REGION Network 7: IW272 - BWT Level (LT-422) - Tank #2
   RUNG wire#powerrail
      { S7_Templates := "[SrcType := Int, DestType := Real]" } Normalize(min := "20_TANKS_IP_DATA".RIO_04.SECOND_TANK.BWT_LEVEL_CNFG.RAW_MIN, value := "Tank 4S BWT Level", max := "20_TANKS_IP_DATA".RIO_04.SECOND_TANK.BWT_LEVEL_CNFG.RAW_MAX, out => "20_TANKS_IP_DATA".RIO_04.SECOND_TANK.BWT_LEVEL_CNFG.NORM)
      { S7_Templates := "[SrcType := Real, DestType := Real]" } Scale(min := "20_TANKS_IP_DATA".RIO_04.SECOND_TANK.BWT_LEVEL_CNFG.ENG_MIN, value := "IN_Level_WBT_4S", max := "20_TANKS_IP_DATA".RIO_04.SECOND_TANK.BWT_LEVEL_CNFG.ENG_MAX, out => "Tag_26")
      Move(in := "Data_From_WBT".Level_WBT_4S, out1 => "20_TANKS_IP_DATA".RIO_04.SECOND_TANK.BWT_LEVEL)
   END_RUNG
   // the same network as SCL:
   "20_TANKS_IP_DATA".RIO_04.SECOND_TANK.BWT_LEVEL_CNFG.NORM := NORM_X(MIN := "20_TANKS_IP_DATA".RIO_04.SECOND_TANK.BWT_LEVEL_CNFG.RAW_MIN, VALUE := "Tank 4S BWT Level", MAX := "20_TANKS_IP_DATA".RIO_04.SECOND_TANK.BWT_LEVEL_CNFG.RAW_MAX);
   "Tag_26" := SCALE_X(MIN := "20_TANKS_IP_DATA".RIO_04.SECOND_TANK.BWT_LEVEL_CNFG.ENG_MIN, VALUE := "IN_Level_WBT_4S", MAX := "20_TANKS_IP_DATA".RIO_04.SECOND_TANK.BWT_LEVEL_CNFG.ENG_MAX);
   "20_TANKS_IP_DATA".RIO_04.SECOND_TANK.BWT_LEVEL := "Data_From_WBT".Level_WBT_4S;
END_REGION

REGION Network 8: IW274 - Spare Input - Tank #1
   RUNG wire#powerrail
      { S7_Templates := "[SrcType := Int, DestType := Real]" } Normalize(min := "20_TANKS_IP_DATA".RIO_04.FIRST_TANK.SPARE_AI_1_CNFG.RAW_MIN, value := "RIO4_SPR_AI_274", max := "20_TANKS_IP_DATA".RIO_04.FIRST_TANK.SPARE_AI_1_CNFG.RAW_MAX, out => "20_TANKS_IP_DATA".RIO_04.FIRST_TANK.SPARE_AI_1_CNFG.NORM)
      { S7_Templates := "[SrcType := Real, DestType := Real]" } Scale(min := "20_TANKS_IP_DATA".RIO_04.FIRST_TANK.SPARE_AI_1_CNFG.ENG_MIN, value := "20_TANKS_IP_DATA".RIO_04.FIRST_TANK.SPARE_AI_1_CNFG.NORM, max := "20_TANKS_IP_DATA".RIO_04.FIRST_TANK.SPARE_AI_1_CNFG.ENG_MAX, out => "20_TANKS_IP_DATA".RIO_04.FIRST_TANK.SPARE_AI_1)
   END_RUNG
   // the same network as SCL:
   "20_TANKS_IP_DATA".RIO_04.FIRST_TANK.SPARE_AI_1_CNFG.NORM := NORM_X(MIN := "20_TANKS_IP_DATA".RIO_04.FIRST_TANK.SPARE_AI_1_CNFG.RAW_MIN, VALUE := "RIO4_SPR_AI_274", MAX := "20_TANKS_IP_DATA".RIO_04.FIRST_TANK.SPARE_AI_1_CNFG.RAW_MAX);
   "20_TANKS_IP_DATA".RIO_04.FIRST_TANK.SPARE_AI_1 := SCALE_X(MIN := "20_TANKS_IP_DATA".RIO_04.FIRST_TANK.SPARE_AI_1_CNFG.ENG_MIN, VALUE := "20_TANKS_IP_DATA".RIO_04.FIRST_TANK.SPARE_AI_1_CNFG.NORM, MAX := "20_TANKS_IP_DATA".RIO_04.FIRST_TANK.SPARE_AI_1_CNFG.ENG_MAX);
END_REGION

REGION Network 9: IW276 - BWT Ph (426) - Tank #1
   RUNG wire#powerrail
      { S7_Templates := "[SrcType := Int, DestType := Real]" } Normalize(min := "20_TANKS_IP_DATA".RIO_04.FIRST_TANK.BWT_PH_CNFG.RAW_MIN, value := "Tank 4P BWT ph", max := "20_TANKS_IP_DATA".RIO_04.FIRST_TANK.BWT_PH_CNFG.RAW_MAX, out => "20_TANKS_IP_DATA".RIO_04.FIRST_TANK.BWT_PH_CNFG.NORM)
      { S7_Templates := "[SrcType := Real, DestType := Real]" } Scale(min := "20_TANKS_IP_DATA".RIO_04.FIRST_TANK.BWT_PH_CNFG.ENG_MIN, value := "20_TANKS_IP_DATA".RIO_04.FIRST_TANK.BWT_PH_CNFG.NORM, max := "20_TANKS_IP_DATA".RIO_04.FIRST_TANK.BWT_PH_CNFG.ENG_MAX, out => "20_TANKS_IP_DATA".RIO_04.FIRST_TANK.BWT_PH)
   END_RUNG
   // the same network as SCL:
   "20_TANKS_IP_DATA".RIO_04.FIRST_TANK.BWT_PH_CNFG.NORM := NORM_X(MIN := "20_TANKS_IP_DATA".RIO_04.FIRST_TANK.BWT_PH_CNFG.RAW_MIN, VALUE := "Tank 4P BWT ph", MAX := "20_TANKS_IP_DATA".RIO_04.FIRST_TANK.BWT_PH_CNFG.RAW_MAX);
   "20_TANKS_IP_DATA".RIO_04.FIRST_TANK.BWT_PH := SCALE_X(MIN := "20_TANKS_IP_DATA".RIO_04.FIRST_TANK.BWT_PH_CNFG.ENG_MIN, VALUE := "20_TANKS_IP_DATA".RIO_04.FIRST_TANK.BWT_PH_CNFG.NORM, MAX := "20_TANKS_IP_DATA".RIO_04.FIRST_TANK.BWT_PH_CNFG.ENG_MAX);
END_REGION

REGION Network 10: IW278 - BWT Temperature (426) - Tank #1
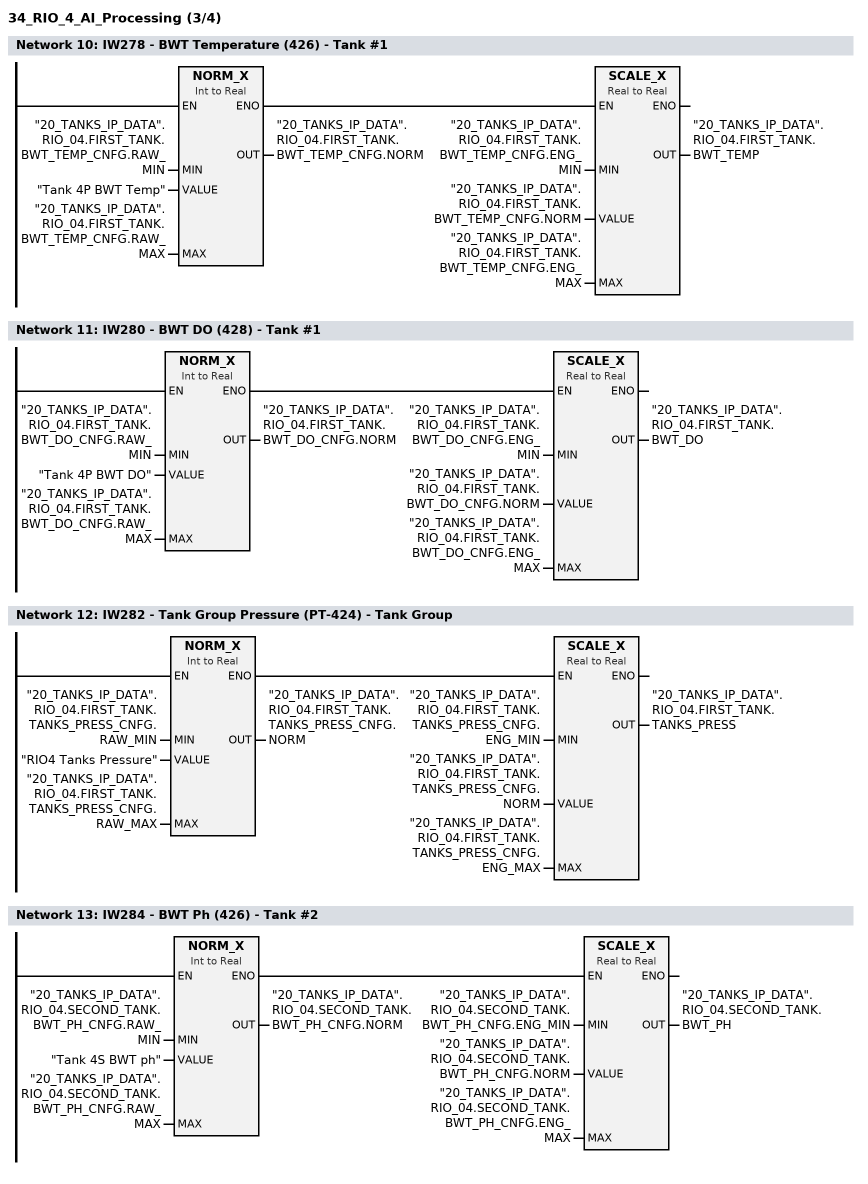
   RUNG wire#powerrail
      { S7_Templates := "[SrcType := Int, DestType := Real]" } Normalize(min := "20_TANKS_IP_DATA".RIO_04.FIRST_TANK.BWT_TEMP_CNFG.RAW_MIN, value := "Tank 4P BWT Temp", max := "20_TANKS_IP_DATA".RIO_04.FIRST_TANK.BWT_TEMP_CNFG.RAW_MAX, out => "20_TANKS_IP_DATA".RIO_04.FIRST_TANK.BWT_TEMP_CNFG.NORM)
      { S7_Templates := "[SrcType := Real, DestType := Real]" } Scale(min := "20_TANKS_IP_DATA".RIO_04.FIRST_TANK.BWT_TEMP_CNFG.ENG_MIN, value := "20_TANKS_IP_DATA".RIO_04.FIRST_TANK.BWT_TEMP_CNFG.NORM, max := "20_TANKS_IP_DATA".RIO_04.FIRST_TANK.BWT_TEMP_CNFG.ENG_MAX, out => "20_TANKS_IP_DATA".RIO_04.FIRST_TANK.BWT_TEMP)
   END_RUNG
   // the same network as SCL:
   "20_TANKS_IP_DATA".RIO_04.FIRST_TANK.BWT_TEMP_CNFG.NORM := NORM_X(MIN := "20_TANKS_IP_DATA".RIO_04.FIRST_TANK.BWT_TEMP_CNFG.RAW_MIN, VALUE := "Tank 4P BWT Temp", MAX := "20_TANKS_IP_DATA".RIO_04.FIRST_TANK.BWT_TEMP_CNFG.RAW_MAX);
   "20_TANKS_IP_DATA".RIO_04.FIRST_TANK.BWT_TEMP := SCALE_X(MIN := "20_TANKS_IP_DATA".RIO_04.FIRST_TANK.BWT_TEMP_CNFG.ENG_MIN, VALUE := "20_TANKS_IP_DATA".RIO_04.FIRST_TANK.BWT_TEMP_CNFG.NORM, MAX := "20_TANKS_IP_DATA".RIO_04.FIRST_TANK.BWT_TEMP_CNFG.ENG_MAX);
END_REGION

REGION Network 11: IW280 - BWT DO (428) - Tank #1
   RUNG wire#powerrail
      { S7_Templates := "[SrcType := Int, DestType := Real]" } Normalize(min := "20_TANKS_IP_DATA".RIO_04.FIRST_TANK.BWT_DO_CNFG.RAW_MIN, value := "Tank 4P BWT DO", max := "20_TANKS_IP_DATA".RIO_04.FIRST_TANK.BWT_DO_CNFG.RAW_MAX, out => "20_TANKS_IP_DATA".RIO_04.FIRST_TANK.BWT_DO_CNFG.NORM)
      { S7_Templates := "[SrcType := Real, DestType := Real]" } Scale(min := "20_TANKS_IP_DATA".RIO_04.FIRST_TANK.BWT_DO_CNFG.ENG_MIN, value := "20_TANKS_IP_DATA".RIO_04.FIRST_TANK.BWT_DO_CNFG.NORM, max := "20_TANKS_IP_DATA".RIO_04.FIRST_TANK.BWT_DO_CNFG.ENG_MAX, out => "20_TANKS_IP_DATA".RIO_04.FIRST_TANK.BWT_DO)
   END_RUNG
   // the same network as SCL:
   "20_TANKS_IP_DATA".RIO_04.FIRST_TANK.BWT_DO_CNFG.NORM := NORM_X(MIN := "20_TANKS_IP_DATA".RIO_04.FIRST_TANK.BWT_DO_CNFG.RAW_MIN, VALUE := "Tank 4P BWT DO", MAX := "20_TANKS_IP_DATA".RIO_04.FIRST_TANK.BWT_DO_CNFG.RAW_MAX);
   "20_TANKS_IP_DATA".RIO_04.FIRST_TANK.BWT_DO := SCALE_X(MIN := "20_TANKS_IP_DATA".RIO_04.FIRST_TANK.BWT_DO_CNFG.ENG_MIN, VALUE := "20_TANKS_IP_DATA".RIO_04.FIRST_TANK.BWT_DO_CNFG.NORM, MAX := "20_TANKS_IP_DATA".RIO_04.FIRST_TANK.BWT_DO_CNFG.ENG_MAX);
END_REGION

REGION Network 12: IW282 - Tank Group Pressure (PT-424) - Tank Group
   RUNG wire#powerrail
      { S7_Templates := "[SrcType := Int, DestType := Real]" } Normalize(min := "20_TANKS_IP_DATA".RIO_04.FIRST_TANK.TANKS_PRESS_CNFG.RAW_MIN, value := "RIO4 Tanks Pressure", max := "20_TANKS_IP_DATA".RIO_04.FIRST_TANK.TANKS_PRESS_CNFG.RAW_MAX, out => "20_TANKS_IP_DATA".RIO_04.FIRST_TANK.TANKS_PRESS_CNFG.NORM)
      { S7_Templates := "[SrcType := Real, DestType := Real]" } Scale(min := "20_TANKS_IP_DATA".RIO_04.FIRST_TANK.TANKS_PRESS_CNFG.ENG_MIN, value := "20_TANKS_IP_DATA".RIO_04.FIRST_TANK.TANKS_PRESS_CNFG.NORM, max := "20_TANKS_IP_DATA".RIO_04.FIRST_TANK.TANKS_PRESS_CNFG.ENG_MAX, out => "20_TANKS_IP_DATA".RIO_04.FIRST_TANK.TANKS_PRESS)
   END_RUNG
   // the same network as SCL:
   "20_TANKS_IP_DATA".RIO_04.FIRST_TANK.TANKS_PRESS_CNFG.NORM := NORM_X(MIN := "20_TANKS_IP_DATA".RIO_04.FIRST_TANK.TANKS_PRESS_CNFG.RAW_MIN, VALUE := "RIO4 Tanks Pressure", MAX := "20_TANKS_IP_DATA".RIO_04.FIRST_TANK.TANKS_PRESS_CNFG.RAW_MAX);
   "20_TANKS_IP_DATA".RIO_04.FIRST_TANK.TANKS_PRESS := SCALE_X(MIN := "20_TANKS_IP_DATA".RIO_04.FIRST_TANK.TANKS_PRESS_CNFG.ENG_MIN, VALUE := "20_TANKS_IP_DATA".RIO_04.FIRST_TANK.TANKS_PRESS_CNFG.NORM, MAX := "20_TANKS_IP_DATA".RIO_04.FIRST_TANK.TANKS_PRESS_CNFG.ENG_MAX);
END_REGION

REGION Network 13: IW284 - BWT Ph (426) - Tank #2
   RUNG wire#powerrail
      { S7_Templates := "[SrcType := Int, DestType := Real]" } Normalize(min := "20_TANKS_IP_DATA".RIO_04.SECOND_TANK.BWT_PH_CNFG.RAW_MIN, value := "Tank 4S BWT ph", max := "20_TANKS_IP_DATA".RIO_04.SECOND_TANK.BWT_PH_CNFG.RAW_MAX, out => "20_TANKS_IP_DATA".RIO_04.SECOND_TANK.BWT_PH_CNFG.NORM)
      { S7_Templates := "[SrcType := Real, DestType := Real]" } Scale(min := "20_TANKS_IP_DATA".RIO_04.SECOND_TANK.BWT_PH_CNFG.ENG_MIN, value := "20_TANKS_IP_DATA".RIO_04.SECOND_TANK.BWT_PH_CNFG.NORM, max := "20_TANKS_IP_DATA".RIO_04.SECOND_TANK.BWT_PH_CNFG.ENG_MAX, out => "20_TANKS_IP_DATA".RIO_04.SECOND_TANK.BWT_PH)
   END_RUNG
   // the same network as SCL:
   "20_TANKS_IP_DATA".RIO_04.SECOND_TANK.BWT_PH_CNFG.NORM := NORM_X(MIN := "20_TANKS_IP_DATA".RIO_04.SECOND_TANK.BWT_PH_CNFG.RAW_MIN, VALUE := "Tank 4S BWT ph", MAX := "20_TANKS_IP_DATA".RIO_04.SECOND_TANK.BWT_PH_CNFG.RAW_MAX);
   "20_TANKS_IP_DATA".RIO_04.SECOND_TANK.BWT_PH := SCALE_X(MIN := "20_TANKS_IP_DATA".RIO_04.SECOND_TANK.BWT_PH_CNFG.ENG_MIN, VALUE := "20_TANKS_IP_DATA".RIO_04.SECOND_TANK.BWT_PH_CNFG.NORM, MAX := "20_TANKS_IP_DATA".RIO_04.SECOND_TANK.BWT_PH_CNFG.ENG_MAX);
END_REGION

REGION Network 14: IW286 - BWT Temperature (426) - Tank #2
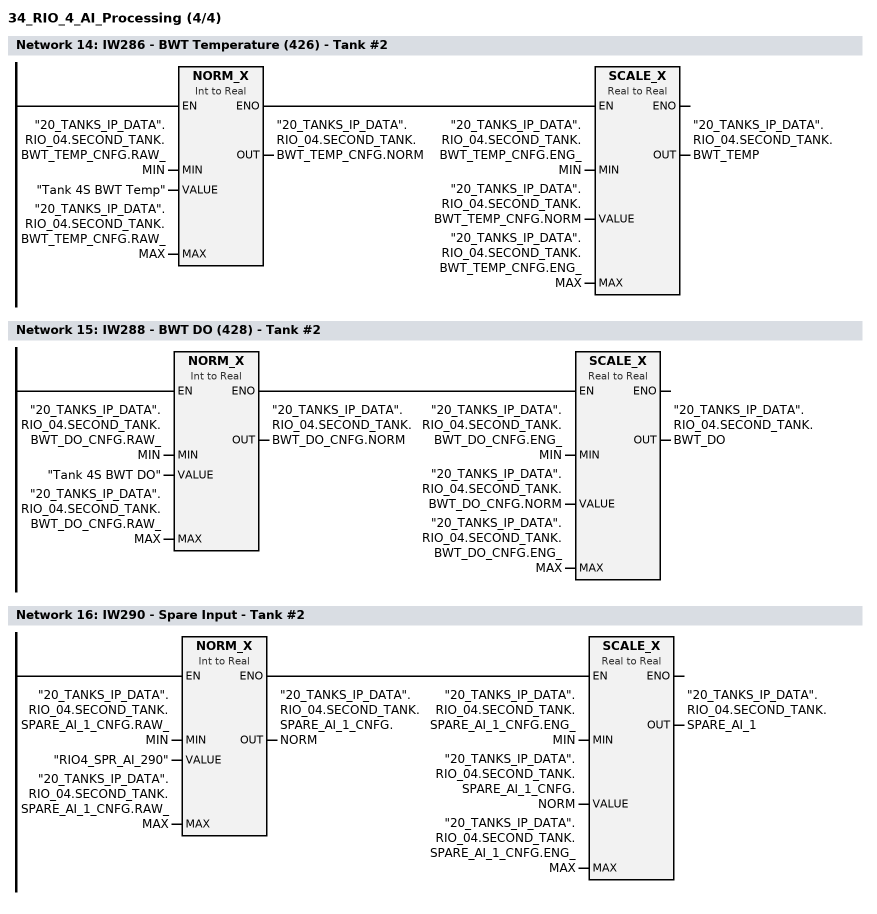
   RUNG wire#powerrail
      { S7_Templates := "[SrcType := Int, DestType := Real]" } Normalize(min := "20_TANKS_IP_DATA".RIO_04.SECOND_TANK.BWT_TEMP_CNFG.RAW_MIN, value := "Tank 4S BWT Temp", max := "20_TANKS_IP_DATA".RIO_04.SECOND_TANK.BWT_TEMP_CNFG.RAW_MAX, out => "20_TANKS_IP_DATA".RIO_04.SECOND_TANK.BWT_TEMP_CNFG.NORM)
      { S7_Templates := "[SrcType := Real, DestType := Real]" } Scale(min := "20_TANKS_IP_DATA".RIO_04.SECOND_TANK.BWT_TEMP_CNFG.ENG_MIN, value := "20_TANKS_IP_DATA".RIO_04.SECOND_TANK.BWT_TEMP_CNFG.NORM, max := "20_TANKS_IP_DATA".RIO_04.SECOND_TANK.BWT_TEMP_CNFG.ENG_MAX, out => "20_TANKS_IP_DATA".RIO_04.SECOND_TANK.BWT_TEMP)
   END_RUNG
   // the same network as SCL:
   "20_TANKS_IP_DATA".RIO_04.SECOND_TANK.BWT_TEMP_CNFG.NORM := NORM_X(MIN := "20_TANKS_IP_DATA".RIO_04.SECOND_TANK.BWT_TEMP_CNFG.RAW_MIN, VALUE := "Tank 4S BWT Temp", MAX := "20_TANKS_IP_DATA".RIO_04.SECOND_TANK.BWT_TEMP_CNFG.RAW_MAX);
   "20_TANKS_IP_DATA".RIO_04.SECOND_TANK.BWT_TEMP := SCALE_X(MIN := "20_TANKS_IP_DATA".RIO_04.SECOND_TANK.BWT_TEMP_CNFG.ENG_MIN, VALUE := "20_TANKS_IP_DATA".RIO_04.SECOND_TANK.BWT_TEMP_CNFG.NORM, MAX := "20_TANKS_IP_DATA".RIO_04.SECOND_TANK.BWT_TEMP_CNFG.ENG_MAX);
END_REGION

REGION Network 15: IW288 - BWT DO (428) - Tank #2
   RUNG wire#powerrail
      { S7_Templates := "[SrcType := Int, DestType := Real]" } Normalize(min := "20_TANKS_IP_DATA".RIO_04.SECOND_TANK.BWT_DO_CNFG.RAW_MIN, value := "Tank 4S BWT DO", max := "20_TANKS_IP_DATA".RIO_04.SECOND_TANK.BWT_DO_CNFG.RAW_MAX, out => "20_TANKS_IP_DATA".RIO_04.SECOND_TANK.BWT_DO_CNFG.NORM)
      { S7_Templates := "[SrcType := Real, DestType := Real]" } Scale(min := "20_TANKS_IP_DATA".RIO_04.SECOND_TANK.BWT_DO_CNFG.ENG_MIN, value := "20_TANKS_IP_DATA".RIO_04.SECOND_TANK.BWT_DO_CNFG.NORM, max := "20_TANKS_IP_DATA".RIO_04.SECOND_TANK.BWT_DO_CNFG.ENG_MAX, out => "20_TANKS_IP_DATA".RIO_04.SECOND_TANK.BWT_DO)
   END_RUNG
   // the same network as SCL:
   "20_TANKS_IP_DATA".RIO_04.SECOND_TANK.BWT_DO_CNFG.NORM := NORM_X(MIN := "20_TANKS_IP_DATA".RIO_04.SECOND_TANK.BWT_DO_CNFG.RAW_MIN, VALUE := "Tank 4S BWT DO", MAX := "20_TANKS_IP_DATA".RIO_04.SECOND_TANK.BWT_DO_CNFG.RAW_MAX);
   "20_TANKS_IP_DATA".RIO_04.SECOND_TANK.BWT_DO := SCALE_X(MIN := "20_TANKS_IP_DATA".RIO_04.SECOND_TANK.BWT_DO_CNFG.ENG_MIN, VALUE := "20_TANKS_IP_DATA".RIO_04.SECOND_TANK.BWT_DO_CNFG.NORM, MAX := "20_TANKS_IP_DATA".RIO_04.SECOND_TANK.BWT_DO_CNFG.ENG_MAX);
END_REGION

REGION Network 16: IW290 - Spare Input - Tank #2
   RUNG wire#powerrail
      { S7_Templates := "[SrcType := Int, DestType := Real]" } Normalize(min := "20_TANKS_IP_DATA".RIO_04.SECOND_TANK.SPARE_AI_1_CNFG.RAW_MIN, value := "RIO4_SPR_AI_290", max := "20_TANKS_IP_DATA".RIO_04.SECOND_TANK.SPARE_AI_1_CNFG.RAW_MAX, out => "20_TANKS_IP_DATA".RIO_04.SECOND_TANK.SPARE_AI_1_CNFG.NORM)
      { S7_Templates := "[SrcType := Real, DestType := Real]" } Scale(min := "20_TANKS_IP_DATA".RIO_04.SECOND_TANK.SPARE_AI_1_CNFG.ENG_MIN, value := "20_TANKS_IP_DATA".RIO_04.SECOND_TANK.SPARE_AI_1_CNFG.NORM, max := "20_TANKS_IP_DATA".RIO_04.SECOND_TANK.SPARE_AI_1_CNFG.ENG_MAX, out => "20_TANKS_IP_DATA".RIO_04.SECOND_TANK.SPARE_AI_1)
   END_RUNG
   // the same network as SCL:
   "20_TANKS_IP_DATA".RIO_04.SECOND_TANK.SPARE_AI_1_CNFG.NORM := NORM_X(MIN := "20_TANKS_IP_DATA".RIO_04.SECOND_TANK.SPARE_AI_1_CNFG.RAW_MIN, VALUE := "RIO4_SPR_AI_290", MAX := "20_TANKS_IP_DATA".RIO_04.SECOND_TANK.SPARE_AI_1_CNFG.RAW_MAX);
   "20_TANKS_IP_DATA".RIO_04.SECOND_TANK.SPARE_AI_1 := SCALE_X(MIN := "20_TANKS_IP_DATA".RIO_04.SECOND_TANK.SPARE_AI_1_CNFG.ENG_MIN, VALUE := "20_TANKS_IP_DATA".RIO_04.SECOND_TANK.SPARE_AI_1_CNFG.NORM, MAX := "20_TANKS_IP_DATA".RIO_04.SECOND_TANK.SPARE_AI_1_CNFG.ENG_MAX);
END_REGION
END_FUNCTION

FUNCTION "35_RIO_5_AI_Processing" : Void   // FC35, LAD
TITLE = Analogue Input Processing (Tank 1 = 5P, Tank 2 = 5S)
{ S7_Optimized_Access := 'TRUE' }
AUTHOR : JRS
VERSION : 0.1
// To process raw inputs prior to code use
BEGIN

REGION Network 1: IW300 - USD Flow (FIT-418) - Tank #1
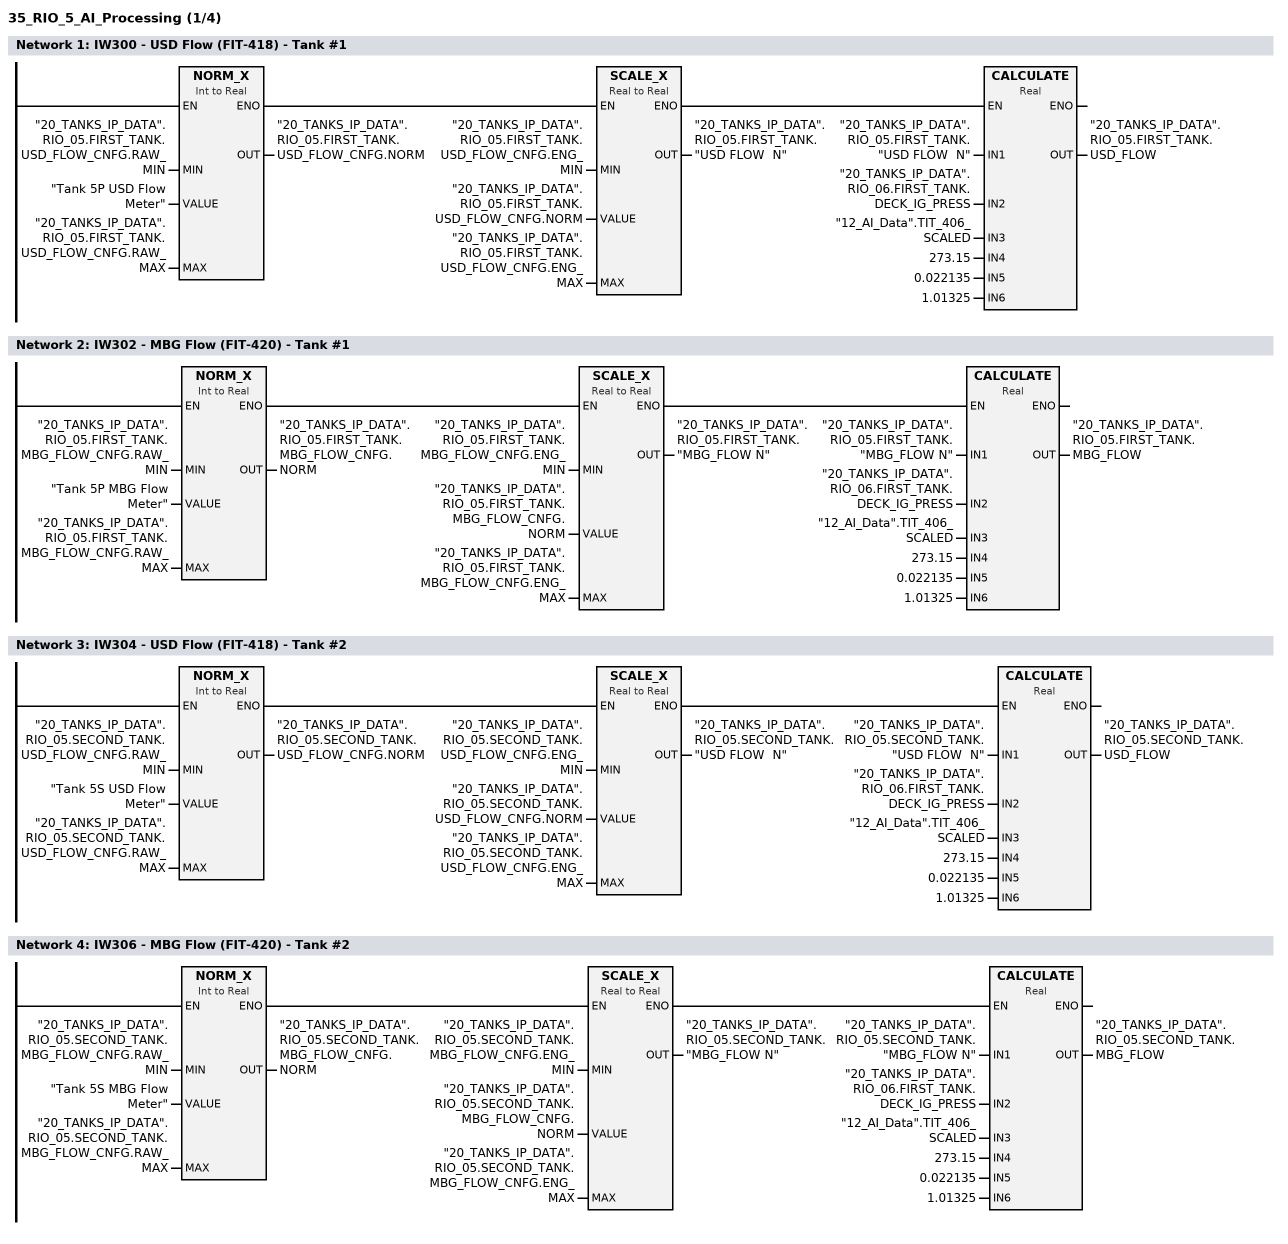
   RUNG wire#powerrail
      { S7_Templates := "[SrcType := Int, DestType := Real]" } Normalize(min := "20_TANKS_IP_DATA".RIO_05.FIRST_TANK.USD_FLOW_CNFG.RAW_MIN, value := "Tank 5P USD Flow Meter", max := "20_TANKS_IP_DATA".RIO_05.FIRST_TANK.USD_FLOW_CNFG.RAW_MAX, out => "20_TANKS_IP_DATA".RIO_05.FIRST_TANK.USD_FLOW_CNFG.NORM)
      { S7_Templates := "[SrcType := Real, DestType := Real]" } Scale(min := "20_TANKS_IP_DATA".RIO_05.FIRST_TANK.USD_FLOW_CNFG.ENG_MIN, value := "20_TANKS_IP_DATA".RIO_05.FIRST_TANK.USD_FLOW_CNFG.NORM, max := "20_TANKS_IP_DATA".RIO_05.FIRST_TANK.USD_FLOW_CNFG.ENG_MAX, out => "20_TANKS_IP_DATA".RIO_05.FIRST_TANK."USD FLOW  N")
      { S7_Templates := "SrcType := Real"; S7_Expression := "IN1*(IN2+IN6)/IN6*IN4/(IN3+IN4)" } Calculate(in1 := "20_TANKS_IP_DATA".RIO_05.FIRST_TANK."USD FLOW  N", in2 := "20_TANKS_IP_DATA".RIO_06.FIRST_TANK.DECK_IG_PRESS, in3 := "12_AI_Data".TIT_406_SCALED, in4 := 273.15, in5 := 0.022135, in6 := 1.01325, out => "20_TANKS_IP_DATA".RIO_05.FIRST_TANK.USD_FLOW)
   END_RUNG
   // the same network as SCL:
   "20_TANKS_IP_DATA".RIO_05.FIRST_TANK.USD_FLOW_CNFG.NORM := NORM_X(MIN := "20_TANKS_IP_DATA".RIO_05.FIRST_TANK.USD_FLOW_CNFG.RAW_MIN, VALUE := "Tank 5P USD Flow Meter", MAX := "20_TANKS_IP_DATA".RIO_05.FIRST_TANK.USD_FLOW_CNFG.RAW_MAX);
   "20_TANKS_IP_DATA".RIO_05.FIRST_TANK."USD FLOW  N" := SCALE_X(MIN := "20_TANKS_IP_DATA".RIO_05.FIRST_TANK.USD_FLOW_CNFG.ENG_MIN, VALUE := "20_TANKS_IP_DATA".RIO_05.FIRST_TANK.USD_FLOW_CNFG.NORM, MAX := "20_TANKS_IP_DATA".RIO_05.FIRST_TANK.USD_FLOW_CNFG.ENG_MAX);
   "20_TANKS_IP_DATA".RIO_05.FIRST_TANK.USD_FLOW := "20_TANKS_IP_DATA".RIO_05.FIRST_TANK."USD FLOW  N"*("20_TANKS_IP_DATA".RIO_06.FIRST_TANK.DECK_IG_PRESS+1.01325)/1.01325*273.15/("12_AI_Data".TIT_406_SCALED+273.15);
END_REGION

REGION Network 2: IW302 - MBG Flow (FIT-420) - Tank #1
   RUNG wire#powerrail
      { S7_Templates := "[SrcType := Int, DestType := Real]" } Normalize(min := "20_TANKS_IP_DATA".RIO_05.FIRST_TANK.MBG_FLOW_CNFG.RAW_MIN, value := "Tank 5P MBG Flow Meter", max := "20_TANKS_IP_DATA".RIO_05.FIRST_TANK.MBG_FLOW_CNFG.RAW_MAX, out => "20_TANKS_IP_DATA".RIO_05.FIRST_TANK.MBG_FLOW_CNFG.NORM)
      { S7_Templates := "[SrcType := Real, DestType := Real]" } Scale(min := "20_TANKS_IP_DATA".RIO_05.FIRST_TANK.MBG_FLOW_CNFG.ENG_MIN, value := "20_TANKS_IP_DATA".RIO_05.FIRST_TANK.MBG_FLOW_CNFG.NORM, max := "20_TANKS_IP_DATA".RIO_05.FIRST_TANK.MBG_FLOW_CNFG.ENG_MAX, out => "20_TANKS_IP_DATA".RIO_05.FIRST_TANK."MBG_FLOW N")
      { S7_Templates := "SrcType := Real"; S7_Expression := "IN1*(IN2+IN6)/IN6*IN4/(IN3+IN4)" } Calculate(in1 := "20_TANKS_IP_DATA".RIO_05.FIRST_TANK."MBG_FLOW N", in2 := "20_TANKS_IP_DATA".RIO_06.FIRST_TANK.DECK_IG_PRESS, in3 := "12_AI_Data".TIT_406_SCALED, in4 := 273.15, in5 := 0.022135, in6 := 1.01325, out => "20_TANKS_IP_DATA".RIO_05.FIRST_TANK.MBG_FLOW)
   END_RUNG
   // the same network as SCL:
   "20_TANKS_IP_DATA".RIO_05.FIRST_TANK.MBG_FLOW_CNFG.NORM := NORM_X(MIN := "20_TANKS_IP_DATA".RIO_05.FIRST_TANK.MBG_FLOW_CNFG.RAW_MIN, VALUE := "Tank 5P MBG Flow Meter", MAX := "20_TANKS_IP_DATA".RIO_05.FIRST_TANK.MBG_FLOW_CNFG.RAW_MAX);
   "20_TANKS_IP_DATA".RIO_05.FIRST_TANK."MBG_FLOW N" := SCALE_X(MIN := "20_TANKS_IP_DATA".RIO_05.FIRST_TANK.MBG_FLOW_CNFG.ENG_MIN, VALUE := "20_TANKS_IP_DATA".RIO_05.FIRST_TANK.MBG_FLOW_CNFG.NORM, MAX := "20_TANKS_IP_DATA".RIO_05.FIRST_TANK.MBG_FLOW_CNFG.ENG_MAX);
   "20_TANKS_IP_DATA".RIO_05.FIRST_TANK.MBG_FLOW := "20_TANKS_IP_DATA".RIO_05.FIRST_TANK."MBG_FLOW N"*("20_TANKS_IP_DATA".RIO_06.FIRST_TANK.DECK_IG_PRESS+1.01325)/1.01325*273.15/("12_AI_Data".TIT_406_SCALED+273.15);
END_REGION

REGION Network 3: IW304 - USD Flow (FIT-418) - Tank #2
   RUNG wire#powerrail
      { S7_Templates := "[SrcType := Int, DestType := Real]" } Normalize(min := "20_TANKS_IP_DATA".RIO_05.SECOND_TANK.USD_FLOW_CNFG.RAW_MIN, value := "Tank 5S USD Flow Meter", max := "20_TANKS_IP_DATA".RIO_05.SECOND_TANK.USD_FLOW_CNFG.RAW_MAX, out => "20_TANKS_IP_DATA".RIO_05.SECOND_TANK.USD_FLOW_CNFG.NORM)
      { S7_Templates := "[SrcType := Real, DestType := Real]" } Scale(min := "20_TANKS_IP_DATA".RIO_05.SECOND_TANK.USD_FLOW_CNFG.ENG_MIN, value := "20_TANKS_IP_DATA".RIO_05.SECOND_TANK.USD_FLOW_CNFG.NORM, max := "20_TANKS_IP_DATA".RIO_05.SECOND_TANK.USD_FLOW_CNFG.ENG_MAX, out => "20_TANKS_IP_DATA".RIO_05.SECOND_TANK."USD FLOW  N")
      { S7_Templates := "SrcType := Real"; S7_Expression := "IN1*(IN2+IN6)/IN6*IN4/(IN3+IN4)" } Calculate(in1 := "20_TANKS_IP_DATA".RIO_05.SECOND_TANK."USD FLOW  N", in2 := "20_TANKS_IP_DATA".RIO_06.FIRST_TANK.DECK_IG_PRESS, in3 := "12_AI_Data".TIT_406_SCALED, in4 := 273.15, in5 := 0.022135, in6 := 1.01325, out => "20_TANKS_IP_DATA".RIO_05.SECOND_TANK.USD_FLOW)
   END_RUNG
   // the same network as SCL:
   "20_TANKS_IP_DATA".RIO_05.SECOND_TANK.USD_FLOW_CNFG.NORM := NORM_X(MIN := "20_TANKS_IP_DATA".RIO_05.SECOND_TANK.USD_FLOW_CNFG.RAW_MIN, VALUE := "Tank 5S USD Flow Meter", MAX := "20_TANKS_IP_DATA".RIO_05.SECOND_TANK.USD_FLOW_CNFG.RAW_MAX);
   "20_TANKS_IP_DATA".RIO_05.SECOND_TANK."USD FLOW  N" := SCALE_X(MIN := "20_TANKS_IP_DATA".RIO_05.SECOND_TANK.USD_FLOW_CNFG.ENG_MIN, VALUE := "20_TANKS_IP_DATA".RIO_05.SECOND_TANK.USD_FLOW_CNFG.NORM, MAX := "20_TANKS_IP_DATA".RIO_05.SECOND_TANK.USD_FLOW_CNFG.ENG_MAX);
   "20_TANKS_IP_DATA".RIO_05.SECOND_TANK.USD_FLOW := "20_TANKS_IP_DATA".RIO_05.SECOND_TANK."USD FLOW  N"*("20_TANKS_IP_DATA".RIO_06.FIRST_TANK.DECK_IG_PRESS+1.01325)/1.01325*273.15/("12_AI_Data".TIT_406_SCALED+273.15);
END_REGION

REGION Network 4: IW306 - MBG Flow (FIT-420) - Tank #2
   RUNG wire#powerrail
      { S7_Templates := "[SrcType := Int, DestType := Real]" } Normalize(min := "20_TANKS_IP_DATA".RIO_05.SECOND_TANK.MBG_FLOW_CNFG.RAW_MIN, value := "Tank 5S MBG Flow Meter", max := "20_TANKS_IP_DATA".RIO_05.SECOND_TANK.MBG_FLOW_CNFG.RAW_MAX, out => "20_TANKS_IP_DATA".RIO_05.SECOND_TANK.MBG_FLOW_CNFG.NORM)
      { S7_Templates := "[SrcType := Real, DestType := Real]" } Scale(min := "20_TANKS_IP_DATA".RIO_05.SECOND_TANK.MBG_FLOW_CNFG.ENG_MIN, value := "20_TANKS_IP_DATA".RIO_05.SECOND_TANK.MBG_FLOW_CNFG.NORM, max := "20_TANKS_IP_DATA".RIO_05.SECOND_TANK.MBG_FLOW_CNFG.ENG_MAX, out => "20_TANKS_IP_DATA".RIO_05.SECOND_TANK."MBG_FLOW N")
      { S7_Templates := "SrcType := Real"; S7_Expression := "IN1*(IN2+IN6)/IN6*IN4/(IN3+IN4)" } Calculate(in1 := "20_TANKS_IP_DATA".RIO_05.SECOND_TANK."MBG_FLOW N", in2 := "20_TANKS_IP_DATA".RIO_06.FIRST_TANK.DECK_IG_PRESS, in3 := "12_AI_Data".TIT_406_SCALED, in4 := 273.15, in5 := 0.022135, in6 := 1.01325, out => "20_TANKS_IP_DATA".RIO_05.SECOND_TANK.MBG_FLOW)
   END_RUNG
   // the same network as SCL:
   "20_TANKS_IP_DATA".RIO_05.SECOND_TANK.MBG_FLOW_CNFG.NORM := NORM_X(MIN := "20_TANKS_IP_DATA".RIO_05.SECOND_TANK.MBG_FLOW_CNFG.RAW_MIN, VALUE := "Tank 5S MBG Flow Meter", MAX := "20_TANKS_IP_DATA".RIO_05.SECOND_TANK.MBG_FLOW_CNFG.RAW_MAX);
   "20_TANKS_IP_DATA".RIO_05.SECOND_TANK."MBG_FLOW N" := SCALE_X(MIN := "20_TANKS_IP_DATA".RIO_05.SECOND_TANK.MBG_FLOW_CNFG.ENG_MIN, VALUE := "20_TANKS_IP_DATA".RIO_05.SECOND_TANK.MBG_FLOW_CNFG.NORM, MAX := "20_TANKS_IP_DATA".RIO_05.SECOND_TANK.MBG_FLOW_CNFG.ENG_MAX);
   "20_TANKS_IP_DATA".RIO_05.SECOND_TANK.MBG_FLOW := "20_TANKS_IP_DATA".RIO_05.SECOND_TANK."MBG_FLOW N"*("20_TANKS_IP_DATA".RIO_06.FIRST_TANK.DECK_IG_PRESS+1.01325)/1.01325*273.15/("12_AI_Data".TIT_406_SCALED+273.15);
END_REGION

REGION Network 5: IW308 - Deck Main IG Pressure (PT-415) - Tank Group
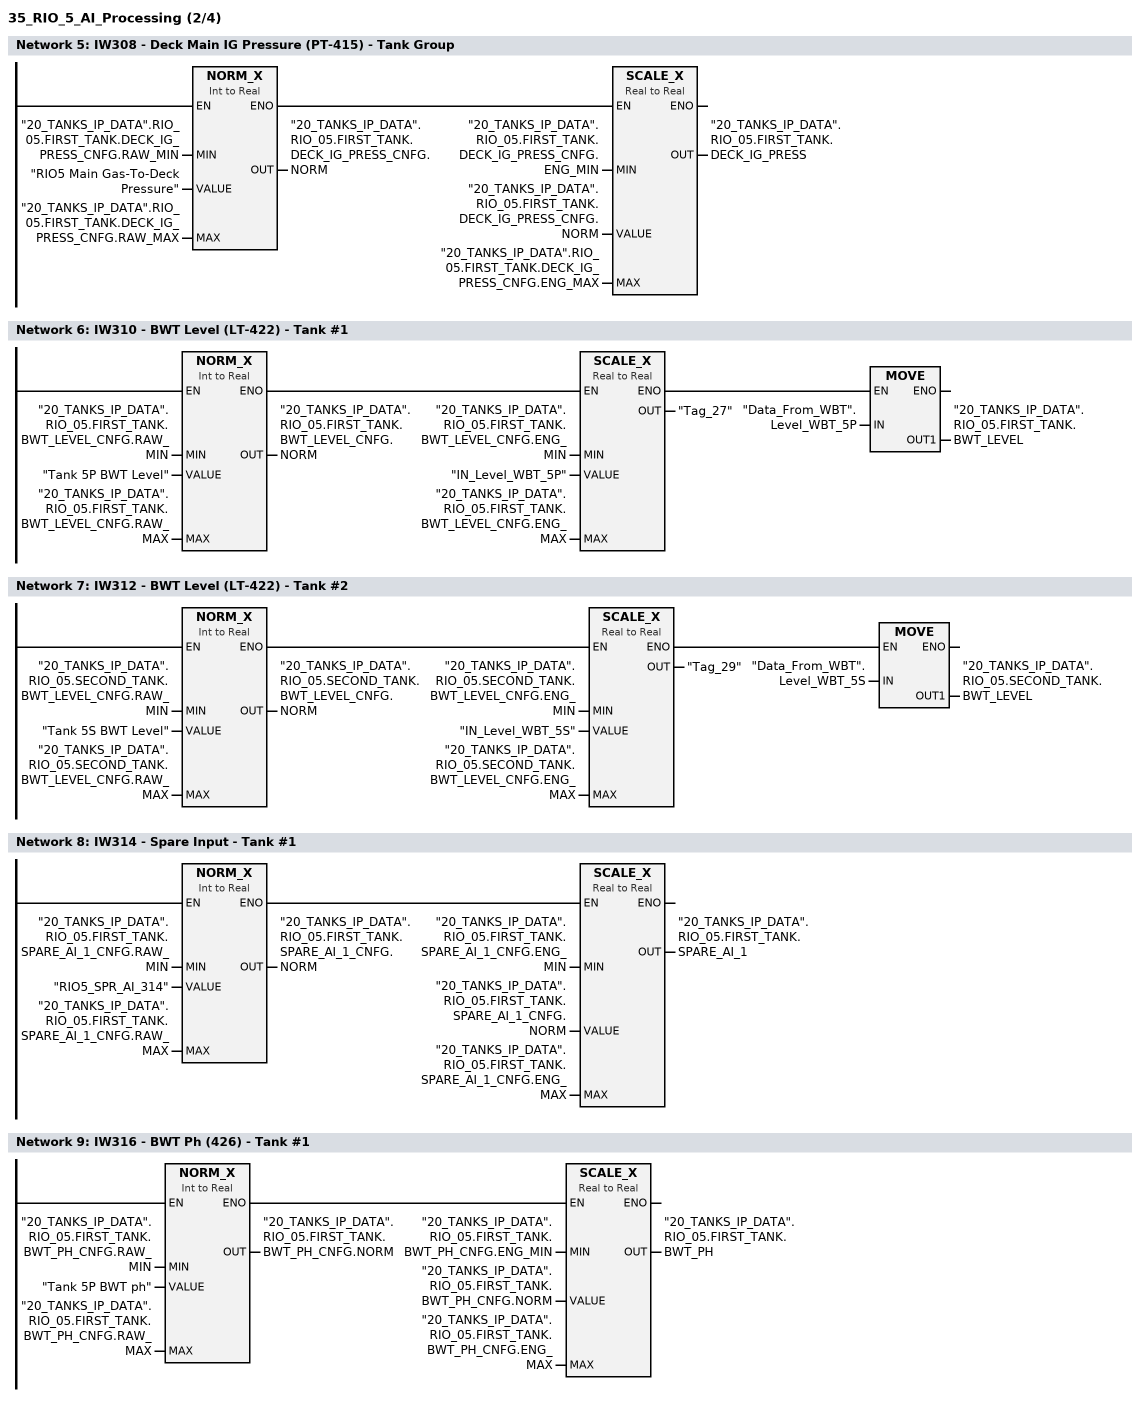
   RUNG wire#powerrail
      { S7_Templates := "[SrcType := Int, DestType := Real]" } Normalize(min := "20_TANKS_IP_DATA".RIO_05.FIRST_TANK.DECK_IG_PRESS_CNFG.RAW_MIN, value := "RIO5 Main Gas-To-Deck Pressure", max := "20_TANKS_IP_DATA".RIO_05.FIRST_TANK.DECK_IG_PRESS_CNFG.RAW_MAX, out => "20_TANKS_IP_DATA".RIO_05.FIRST_TANK.DECK_IG_PRESS_CNFG.NORM)
      { S7_Templates := "[SrcType := Real, DestType := Real]" } Scale(min := "20_TANKS_IP_DATA".RIO_05.FIRST_TANK.DECK_IG_PRESS_CNFG.ENG_MIN, value := "20_TANKS_IP_DATA".RIO_05.FIRST_TANK.DECK_IG_PRESS_CNFG.NORM, max := "20_TANKS_IP_DATA".RIO_05.FIRST_TANK.DECK_IG_PRESS_CNFG.ENG_MAX, out => "20_TANKS_IP_DATA".RIO_05.FIRST_TANK.DECK_IG_PRESS)
   END_RUNG
   // the same network as SCL:
   "20_TANKS_IP_DATA".RIO_05.FIRST_TANK.DECK_IG_PRESS_CNFG.NORM := NORM_X(MIN := "20_TANKS_IP_DATA".RIO_05.FIRST_TANK.DECK_IG_PRESS_CNFG.RAW_MIN, VALUE := "RIO5 Main Gas-To-Deck Pressure", MAX := "20_TANKS_IP_DATA".RIO_05.FIRST_TANK.DECK_IG_PRESS_CNFG.RAW_MAX);
   "20_TANKS_IP_DATA".RIO_05.FIRST_TANK.DECK_IG_PRESS := SCALE_X(MIN := "20_TANKS_IP_DATA".RIO_05.FIRST_TANK.DECK_IG_PRESS_CNFG.ENG_MIN, VALUE := "20_TANKS_IP_DATA".RIO_05.FIRST_TANK.DECK_IG_PRESS_CNFG.NORM, MAX := "20_TANKS_IP_DATA".RIO_05.FIRST_TANK.DECK_IG_PRESS_CNFG.ENG_MAX);
END_REGION

REGION Network 6: IW310 - BWT Level (LT-422) - Tank #1
   RUNG wire#powerrail
      { S7_Templates := "[SrcType := Int, DestType := Real]" } Normalize(min := "20_TANKS_IP_DATA".RIO_05.FIRST_TANK.BWT_LEVEL_CNFG.RAW_MIN, value := "Tank 5P BWT Level", max := "20_TANKS_IP_DATA".RIO_05.FIRST_TANK.BWT_LEVEL_CNFG.RAW_MAX, out => "20_TANKS_IP_DATA".RIO_05.FIRST_TANK.BWT_LEVEL_CNFG.NORM)
      { S7_Templates := "[SrcType := Real, DestType := Real]" } Scale(min := "20_TANKS_IP_DATA".RIO_05.FIRST_TANK.BWT_LEVEL_CNFG.ENG_MIN, value := "IN_Level_WBT_5P", max := "20_TANKS_IP_DATA".RIO_05.FIRST_TANK.BWT_LEVEL_CNFG.ENG_MAX, out => "Tag_27")
      Move(in := "Data_From_WBT".Level_WBT_5P, out1 => "20_TANKS_IP_DATA".RIO_05.FIRST_TANK.BWT_LEVEL)
   END_RUNG
   // the same network as SCL:
   "20_TANKS_IP_DATA".RIO_05.FIRST_TANK.BWT_LEVEL_CNFG.NORM := NORM_X(MIN := "20_TANKS_IP_DATA".RIO_05.FIRST_TANK.BWT_LEVEL_CNFG.RAW_MIN, VALUE := "Tank 5P BWT Level", MAX := "20_TANKS_IP_DATA".RIO_05.FIRST_TANK.BWT_LEVEL_CNFG.RAW_MAX);
   "Tag_27" := SCALE_X(MIN := "20_TANKS_IP_DATA".RIO_05.FIRST_TANK.BWT_LEVEL_CNFG.ENG_MIN, VALUE := "IN_Level_WBT_5P", MAX := "20_TANKS_IP_DATA".RIO_05.FIRST_TANK.BWT_LEVEL_CNFG.ENG_MAX);
   "20_TANKS_IP_DATA".RIO_05.FIRST_TANK.BWT_LEVEL := "Data_From_WBT".Level_WBT_5P;
END_REGION

REGION Network 7: IW312 - BWT Level (LT-422) - Tank #2
   RUNG wire#powerrail
      { S7_Templates := "[SrcType := Int, DestType := Real]" } Normalize(min := "20_TANKS_IP_DATA".RIO_05.SECOND_TANK.BWT_LEVEL_CNFG.RAW_MIN, value := "Tank 5S BWT Level", max := "20_TANKS_IP_DATA".RIO_05.SECOND_TANK.BWT_LEVEL_CNFG.RAW_MAX, out => "20_TANKS_IP_DATA".RIO_05.SECOND_TANK.BWT_LEVEL_CNFG.NORM)
      { S7_Templates := "[SrcType := Real, DestType := Real]" } Scale(min := "20_TANKS_IP_DATA".RIO_05.SECOND_TANK.BWT_LEVEL_CNFG.ENG_MIN, value := "IN_Level_WBT_5S", max := "20_TANKS_IP_DATA".RIO_05.SECOND_TANK.BWT_LEVEL_CNFG.ENG_MAX, out => "Tag_29")
      Move(in := "Data_From_WBT".Level_WBT_5S, out1 => "20_TANKS_IP_DATA".RIO_05.SECOND_TANK.BWT_LEVEL)
   END_RUNG
   // the same network as SCL:
   "20_TANKS_IP_DATA".RIO_05.SECOND_TANK.BWT_LEVEL_CNFG.NORM := NORM_X(MIN := "20_TANKS_IP_DATA".RIO_05.SECOND_TANK.BWT_LEVEL_CNFG.RAW_MIN, VALUE := "Tank 5S BWT Level", MAX := "20_TANKS_IP_DATA".RIO_05.SECOND_TANK.BWT_LEVEL_CNFG.RAW_MAX);
   "Tag_29" := SCALE_X(MIN := "20_TANKS_IP_DATA".RIO_05.SECOND_TANK.BWT_LEVEL_CNFG.ENG_MIN, VALUE := "IN_Level_WBT_5S", MAX := "20_TANKS_IP_DATA".RIO_05.SECOND_TANK.BWT_LEVEL_CNFG.ENG_MAX);
   "20_TANKS_IP_DATA".RIO_05.SECOND_TANK.BWT_LEVEL := "Data_From_WBT".Level_WBT_5S;
END_REGION
